(* Logix 5000 project; controller _GigaDiscovery vendor 1 type 14 code 244 rev 35.11; software revision 35.03; part 12 of 23 *)
(* tags used below, declared in another part *)
   LapBars_Alarms_Time : DINT;
   Timer : TIMER[60];
   Timer_Restraints_Open : TIMER[41];
   DC_Field_Motor_7 : UDT_CROUT;   // DC Field Motor 7 Gondola Contactor -Q16101E -Q16103E
   DC_Field_Pylon_Motors : UDT_CROUT;   // DC Field Pylon Motors Contactor -Q10101E -Q10103E
   Emergencies_CL1 : DINT[14];
   Gondola_Drive_Enable : UDT_CROUT;   // Gondola Drive Ch1-Ch2 Start Enable Contactors -Q16105E -Q16107E
   I_EStop_Pb_OCC1 : UDT_DCI_STOP_TEST;   // +OCC E-stop -S30301F
   I_EStop_Pb_OCC2 : UDT_DCI_STOP_TEST;   // +OCC2 E-Stop -S28502F
   I_OCC2_ACONFIRM : BOOL;   // OCC2 Allow Main CONFIRM -S28602F
   I_OCC2_Disable : UDT_DCM;   // OCC 2 CONTROL DISABLE Page 310
   I_OCC2_RESTRAINTS_RELEASE : Sel_3_Pos_2_Input;   // -S28507F RESTRAINTS RELEASE UNLOCK -RUN- LOCK
   I_OCC_Aut_Man_Selector_Motion : UDT_DCM;   // S30801F
   I_OCC_LockOut_Motion : UDT_DCM;   // OCC -Lockout Motion -Q31203E
   I_OCC_Memory_Footpedal : BOOL;
   I_OCC_Temperature_OK : BOOL;   // OCC temperature OK -S31003E
   I_RESTRAINTS_Selector : Sel_3_Pos_2_Input;   // RESTRAINTS Selctor -S30505F Left = Open Right = Close Center = Nothing
   I_Start_PB : Start_AOI;   // Primary console Strat Push botton Right and Left -S30401F -S30403F
   No_Sfty : Std_to_Sfty;
   O_RESTRAINTS_MainValve : UDT_CROUT;   // Main Valve -B40501I
   Power_On_Delay : BOOL;
   Pylon_Start_Drive_1_2 : UDT_CROUT;   // Pylon Start Drive 1 - 2 Contactors -Q9002H -Q9004H -Q10202G
   Pylon_Start_Drive_3_4 : UDT_CROUT;   // Pylon Start Drive 3 - 4 Contactors -Q9005H -Q9007H -Q12202G
   Pylon_Start_Drive_5_6 : UDT_CROUT;   // Pylon Start Drive 5 - 6 Contactors -Q9009E -Q9011E4 -Q14202G -Q14202G
   RESTRAINTS_MainValve_PressTest : Valve_2_pos_monostable;
   RESTRAINTS_Sector : LapBars_Sector[9];
   Start_Stop_Cycle : Sequencer;
(* S_Alarms, continued *)

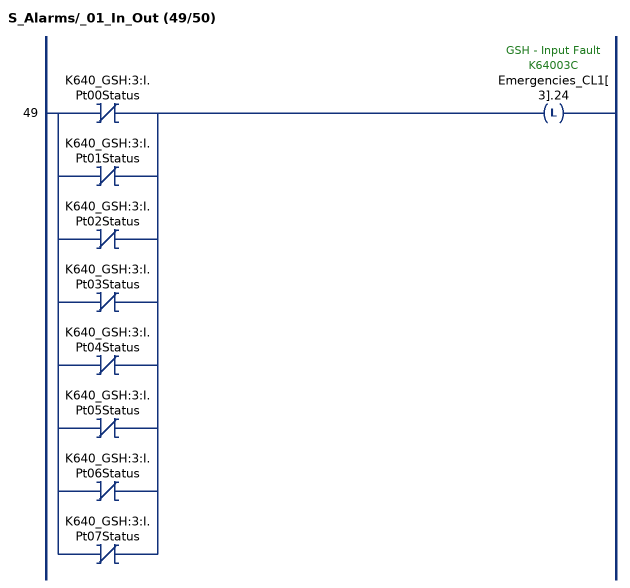
   [picture p209: S_Alarms/_01_In_Out rungs 49-49]
   49: [XIO(K640_GSH:3:I.Pt00Status) ,XIO(K640_GSH:3:I.Pt01Status) ,XIO(K640_GSH:3:I.Pt02Status) ,XIO(K640_GSH:3:I.Pt03Status) ,XIO(K640_GSH:3:I.Pt04Status) ,XIO(K640_GSH:3:I.Pt05Status) ,XIO(K640_GSH:3:I.Pt06Status) ,XIO(K640_GSH:3:I.Pt07Status) ]OTL(Emergencies_CL1[3].24);
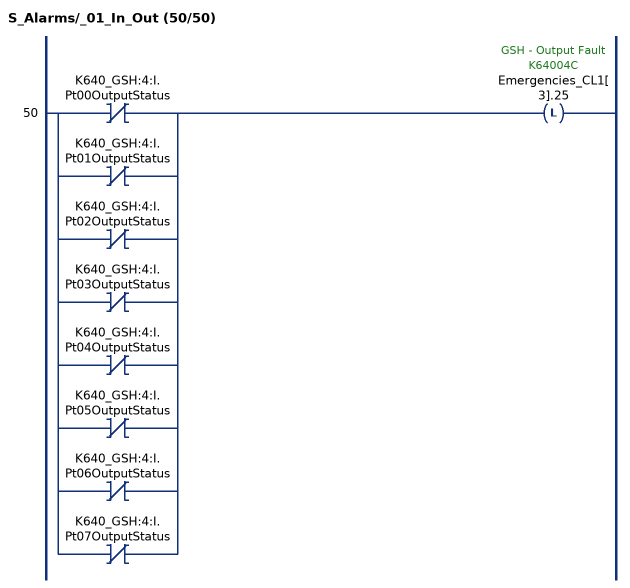
   50: [XIO(K640_GSH:4:I.Pt00OutputStatus) ,XIO(K640_GSH:4:I.Pt01OutputStatus) ,XIO(K640_GSH:4:I.Pt02OutputStatus) ,XIO(K640_GSH:4:I.Pt03OutputStatus) ,XIO(K640_GSH:4:I.Pt04OutputStatus) ,XIO(K640_GSH:4:I.Pt05OutputStatus) ,XIO(K640_GSH:4:I.Pt06OutputStatus) ,XIO(K640_GSH:4:I.Pt07OutputStatus) ]OTL(Emergencies_CL1[3].25);
END_ROUTINE

ROUTINE _02_OCCs   (* ladder *)
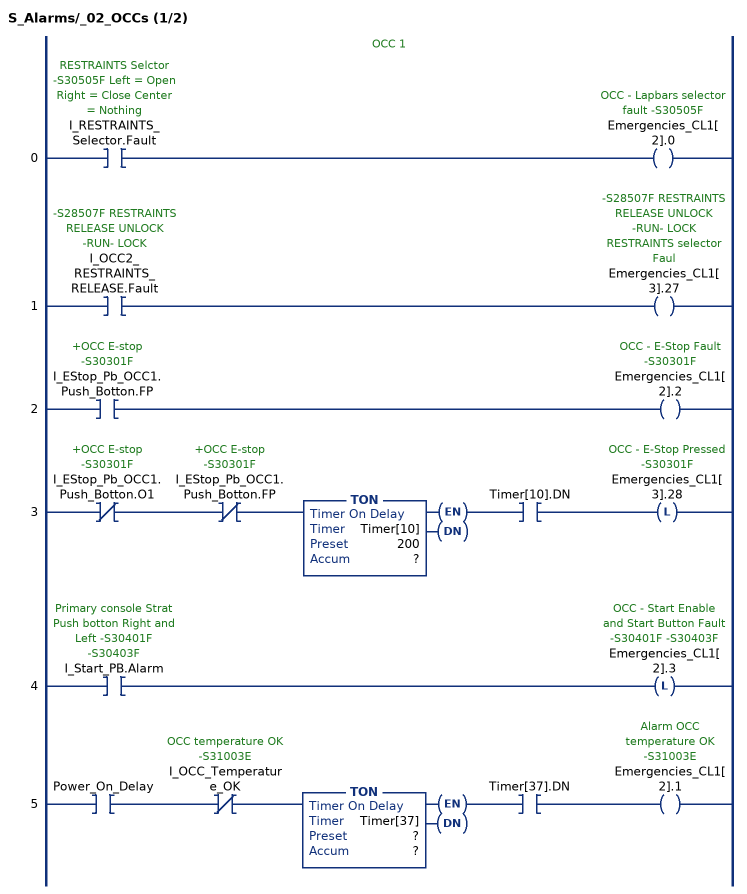
   // OCC 1
   0: XIC(I_RESTRAINTS_Selector.Fault)OTE(Emergencies_CL1[2].0);
   1: XIC(I_OCC2_RESTRAINTS_RELEASE.Fault)OTE(Emergencies_CL1[3].27);
   2: XIC(I_EStop_Pb_OCC1.Push_Botton.FP)OTE(Emergencies_CL1[2].2);
   3: XIO(I_EStop_Pb_OCC1.Push_Botton.O1)XIO(I_EStop_Pb_OCC1.Push_Botton.FP)TON(Timer[10],?,?)XIC(Timer[10].DN)OTL(Emergencies_CL1[3].28);
   4: XIC(I_Start_PB.Alarm)OTL(Emergencies_CL1[2].3);
   5: XIC(Power_On_Delay)XIO(I_OCC_Temperature_OK)TON(Timer[37],?,?)XIC(Timer[37].DN)OTE(Emergencies_CL1[2].1);
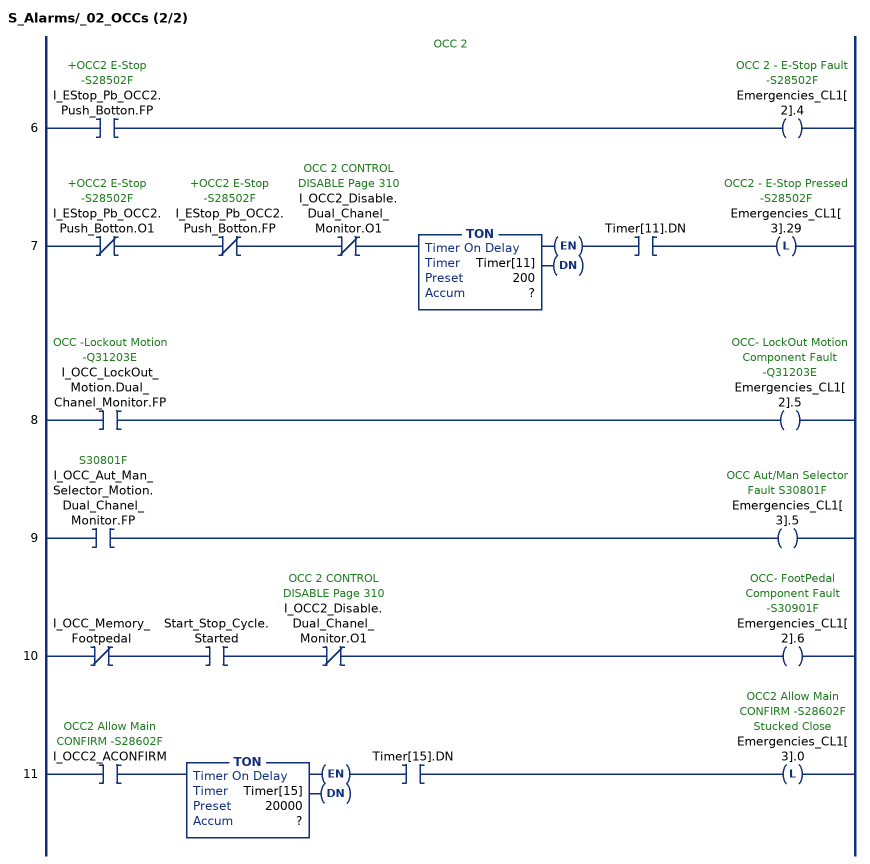
   // OCC 2
   6: XIC(I_EStop_Pb_OCC2.Push_Botton.FP)OTE(Emergencies_CL1[2].4);
   7: XIO(I_EStop_Pb_OCC2.Push_Botton.O1)XIO(I_EStop_Pb_OCC2.Push_Botton.FP)XIO(I_OCC2_Disable.Dual_Chanel_Monitor.O1)TON(Timer[11],?,?)XIC(Timer[11].DN)OTL(Emergencies_CL1[3].29);
   8: XIC(I_OCC_LockOut_Motion.Dual_Chanel_Monitor.FP)OTE(Emergencies_CL1[2].5);
   9: XIC(I_OCC_Aut_Man_Selector_Motion.Dual_Chanel_Monitor.FP)OTE(Emergencies_CL1[3].5);
   10: XIO(I_OCC_Memory_Footpedal)XIC(Start_Stop_Cycle.Started)XIO(I_OCC2_Disable.Dual_Chanel_Monitor.O1)OTE(Emergencies_CL1[2].6);
   11: XIC(I_OCC2_ACONFIRM)TON(Timer[15],?,?)XIC(Timer[15].DN)OTL(Emergencies_CL1[3].0);
END_ROUTINE

ROUTINE _03_MCC   (* ladder *)
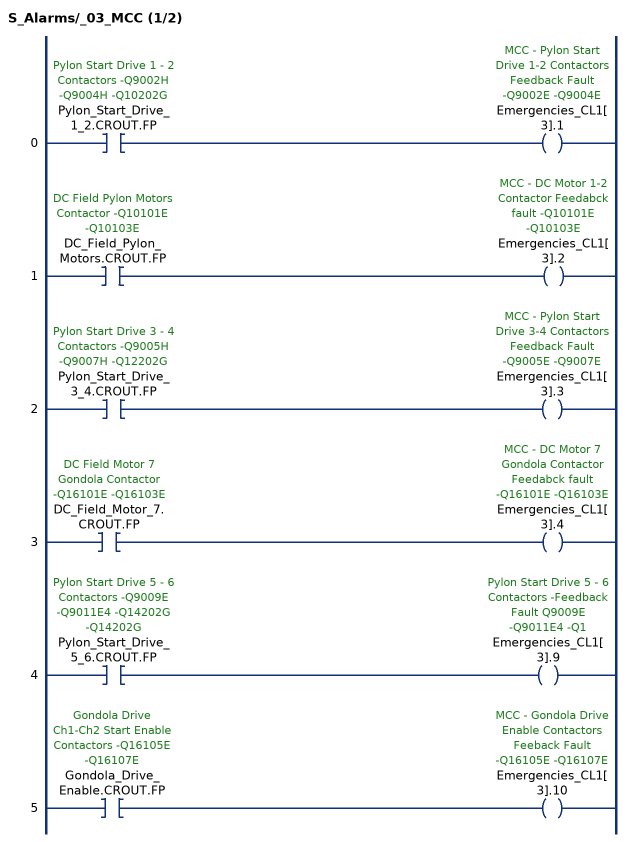
   0: XIC(Pylon_Start_Drive_1_2.CROUT.FP)OTE(Emergencies_CL1[3].1);
   1: XIC(DC_Field_Pylon_Motors.CROUT.FP)OTE(Emergencies_CL1[3].2);
   2: XIC(Pylon_Start_Drive_3_4.CROUT.FP)OTE(Emergencies_CL1[3].3);
   3: XIC(DC_Field_Motor_7.CROUT.FP)OTE(Emergencies_CL1[3].4);
   4: XIC(Pylon_Start_Drive_5_6.CROUT.FP)OTE(Emergencies_CL1[3].9);
   5: XIC(Gondola_Drive_Enable.CROUT.FP)OTE(Emergencies_CL1[3].10);
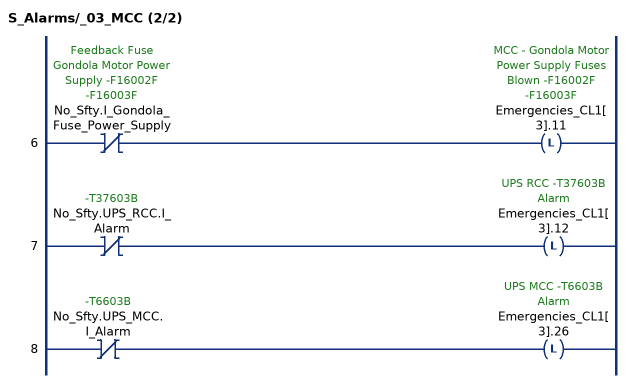
   6: XIO(No_Sfty.I_Gondola_Fuse_Power_Supply)OTL(Emergencies_CL1[3].11);
   7: XIO(No_Sfty.UPS_RCC.I_Alarm)OTL(Emergencies_CL1[3].12);
   8: XIO(No_Sfty.UPS_MCC.I_Alarm)OTL(Emergencies_CL1[3].26);
END_ROUTINE

ROUTINE _04_RESTRAINT_RELEASE   (* ladder *)
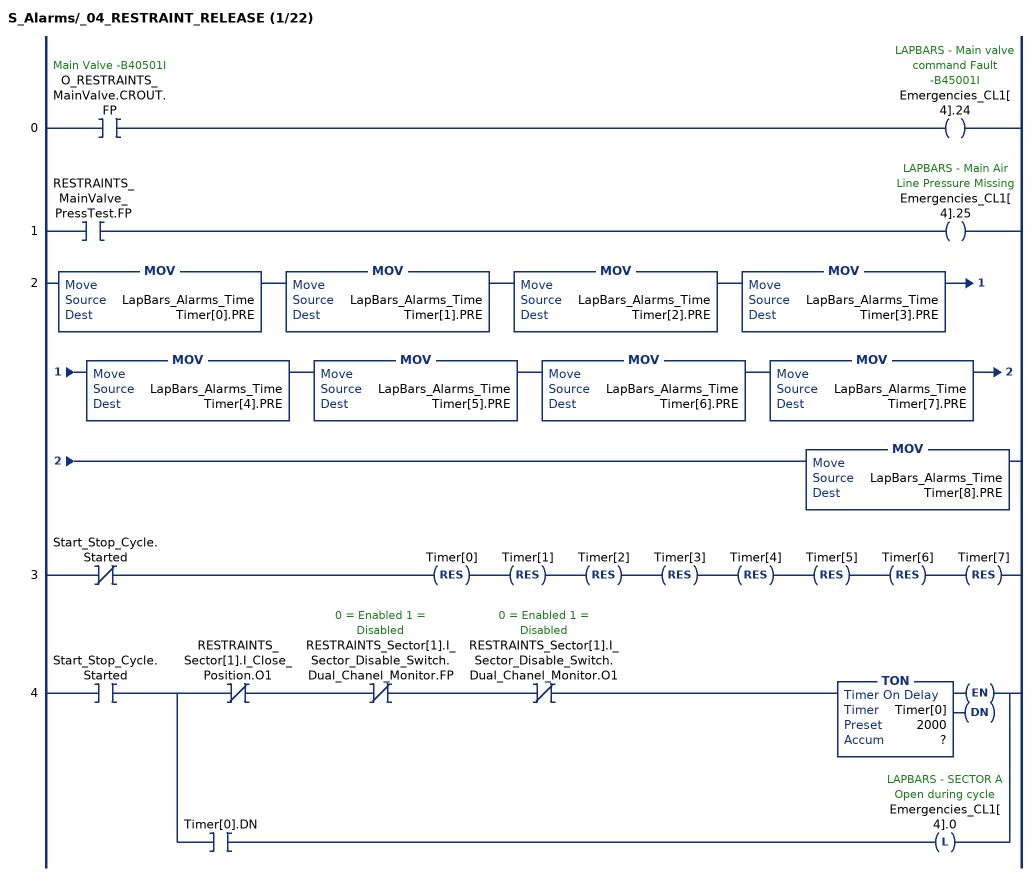
   0: XIC(O_RESTRAINTS_MainValve.CROUT.FP)OTE(Emergencies_CL1[4].24);
   1: XIC(RESTRAINTS_MainValve_PressTest.FP)OTE(Emergencies_CL1[4].25);
   2: MOV(LapBars_Alarms_Time,Timer[0].PRE)MOV(LapBars_Alarms_Time,Timer[1].PRE)MOV(LapBars_Alarms_Time,Timer[2].PRE)MOV(LapBars_Alarms_Time,Timer[3].PRE)MOV(LapBars_Alarms_Time,Timer[4].PRE)MOV(LapBars_Alarms_Time,Timer[5].PRE)MOV(LapBars_Alarms_Time,Timer[6].PRE)MOV(LapBars_Alarms_Time,Timer[7].PRE)MOV(LapBars_Alarms_Time,Timer[8].PRE);
   3: XIO(Start_Stop_Cycle.Started)RES(Timer[0])RES(Timer[1])RES(Timer[2])RES(Timer[3])RES(Timer[4])RES(Timer[5])RES(Timer[6])RES(Timer[7]);
   4: XIC(Start_Stop_Cycle.Started)[XIO(RESTRAINTS_Sector[1].I_Close_Position.O1) XIO(RESTRAINTS_Sector[1].I_Sector_Disable_Switch.Dual_Chanel_Monitor.FP) XIO(RESTRAINTS_Sector[1].I_Sector_Disable_Switch.Dual_Chanel_Monitor.O1) TON(Timer[0],?,?) ,XIC(Timer[0].DN) OTL(Emergencies_CL1[4].0) ];
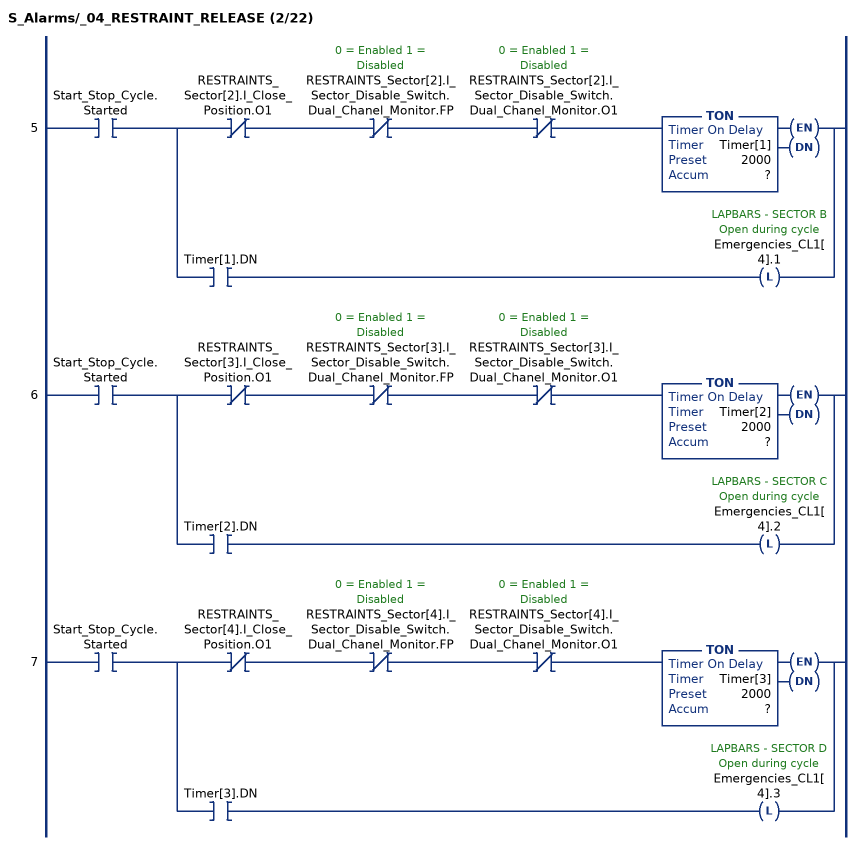
   5: XIC(Start_Stop_Cycle.Started)[XIO(RESTRAINTS_Sector[2].I_Close_Position.O1) XIO(RESTRAINTS_Sector[2].I_Sector_Disable_Switch.Dual_Chanel_Monitor.FP) XIO(RESTRAINTS_Sector[2].I_Sector_Disable_Switch.Dual_Chanel_Monitor.O1) TON(Timer[1],?,?) ,XIC(Timer[1].DN) OTL(Emergencies_CL1[4].1) ];
   6: XIC(Start_Stop_Cycle.Started)[XIO(RESTRAINTS_Sector[3].I_Close_Position.O1) XIO(RESTRAINTS_Sector[3].I_Sector_Disable_Switch.Dual_Chanel_Monitor.FP) XIO(RESTRAINTS_Sector[3].I_Sector_Disable_Switch.Dual_Chanel_Monitor.O1) TON(Timer[2],?,?) ,XIC(Timer[2].DN) OTL(Emergencies_CL1[4].2) ];
   7: XIC(Start_Stop_Cycle.Started)[XIO(RESTRAINTS_Sector[4].I_Close_Position.O1) XIO(RESTRAINTS_Sector[4].I_Sector_Disable_Switch.Dual_Chanel_Monitor.FP) XIO(RESTRAINTS_Sector[4].I_Sector_Disable_Switch.Dual_Chanel_Monitor.O1) TON(Timer[3],?,?) ,XIC(Timer[3].DN) OTL(Emergencies_CL1[4].3) ];
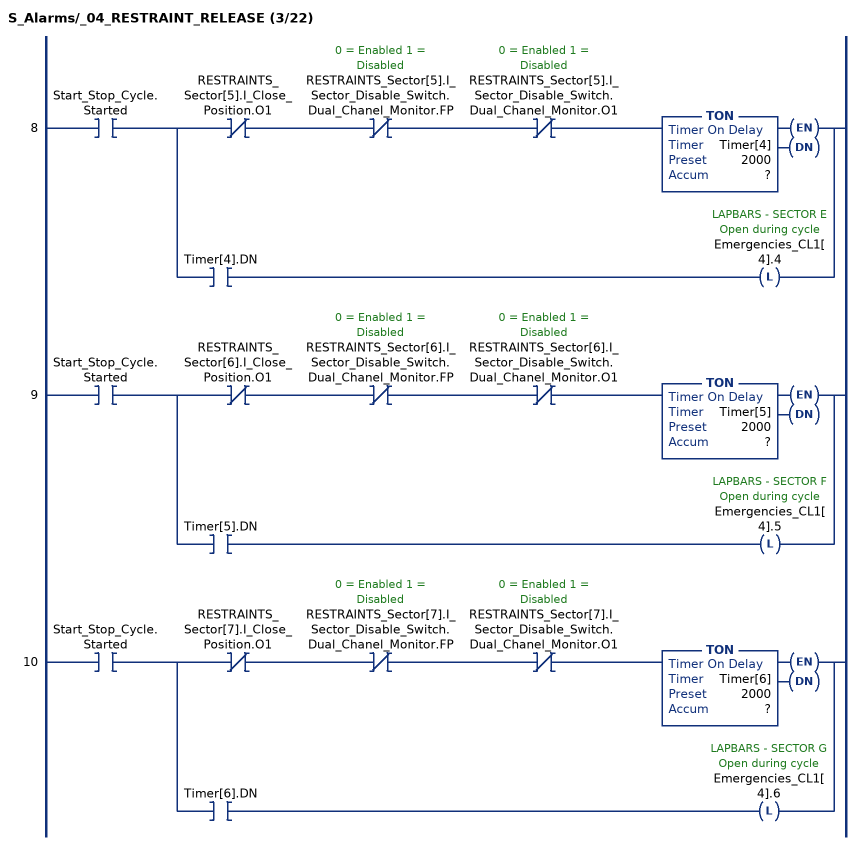
   8: XIC(Start_Stop_Cycle.Started)[XIO(RESTRAINTS_Sector[5].I_Close_Position.O1) XIO(RESTRAINTS_Sector[5].I_Sector_Disable_Switch.Dual_Chanel_Monitor.FP) XIO(RESTRAINTS_Sector[5].I_Sector_Disable_Switch.Dual_Chanel_Monitor.O1) TON(Timer[4],?,?) ,XIC(Timer[4].DN) OTL(Emergencies_CL1[4].4) ];
   9: XIC(Start_Stop_Cycle.Started)[XIO(RESTRAINTS_Sector[6].I_Close_Position.O1) XIO(RESTRAINTS_Sector[6].I_Sector_Disable_Switch.Dual_Chanel_Monitor.FP) XIO(RESTRAINTS_Sector[6].I_Sector_Disable_Switch.Dual_Chanel_Monitor.O1) TON(Timer[5],?,?) ,XIC(Timer[5].DN) OTL(Emergencies_CL1[4].5) ];
   10: XIC(Start_Stop_Cycle.Started)[XIO(RESTRAINTS_Sector[7].I_Close_Position.O1) XIO(RESTRAINTS_Sector[7].I_Sector_Disable_Switch.Dual_Chanel_Monitor.FP) XIO(RESTRAINTS_Sector[7].I_Sector_Disable_Switch.Dual_Chanel_Monitor.O1) TON(Timer[6],?,?) ,XIC(Timer[6].DN) OTL(Emergencies_CL1[4].6) ];
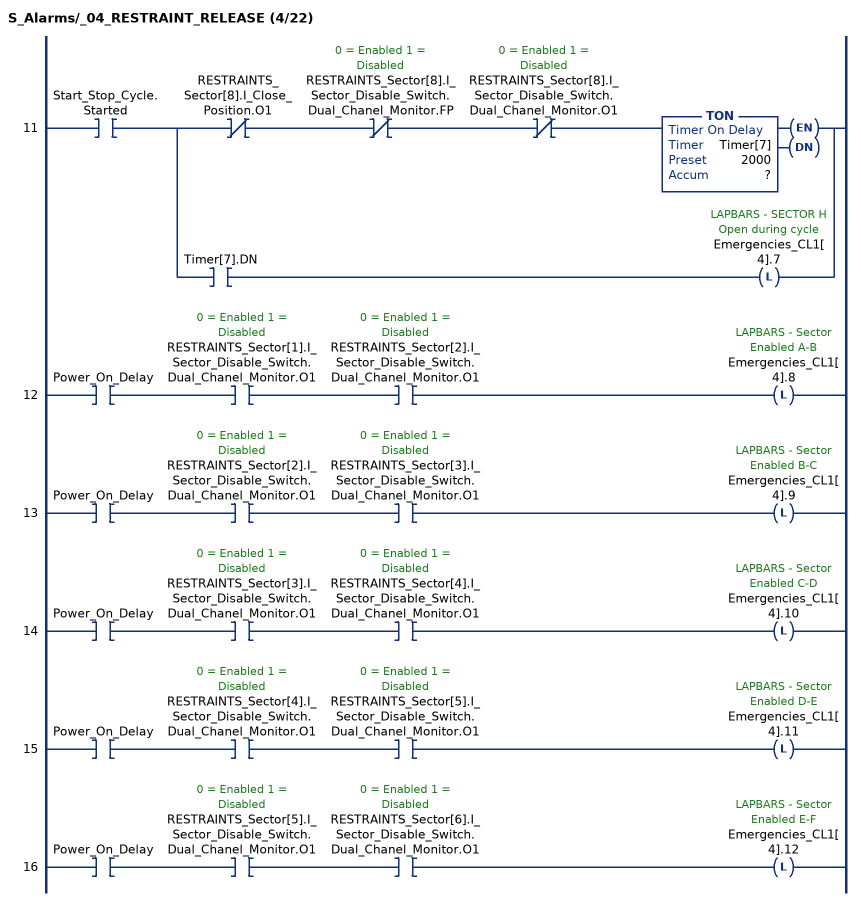
   11: XIC(Start_Stop_Cycle.Started)[XIO(RESTRAINTS_Sector[8].I_Close_Position.O1) XIO(RESTRAINTS_Sector[8].I_Sector_Disable_Switch.Dual_Chanel_Monitor.FP) XIO(RESTRAINTS_Sector[8].I_Sector_Disable_Switch.Dual_Chanel_Monitor.O1) TON(Timer[7],?,?) ,XIC(Timer[7].DN) OTL(Emergencies_CL1[4].7) ];
   12: XIC(Power_On_Delay)XIC(RESTRAINTS_Sector[1].I_Sector_Disable_Switch.Dual_Chanel_Monitor.O1)XIC(RESTRAINTS_Sector[2].I_Sector_Disable_Switch.Dual_Chanel_Monitor.O1)OTL(Emergencies_CL1[4].8);
   13: XIC(Power_On_Delay)XIC(RESTRAINTS_Sector[2].I_Sector_Disable_Switch.Dual_Chanel_Monitor.O1)XIC(RESTRAINTS_Sector[3].I_Sector_Disable_Switch.Dual_Chanel_Monitor.O1)OTL(Emergencies_CL1[4].9);
   14: XIC(Power_On_Delay)XIC(RESTRAINTS_Sector[3].I_Sector_Disable_Switch.Dual_Chanel_Monitor.O1)XIC(RESTRAINTS_Sector[4].I_Sector_Disable_Switch.Dual_Chanel_Monitor.O1)OTL(Emergencies_CL1[4].10);
   15: XIC(Power_On_Delay)XIC(RESTRAINTS_Sector[4].I_Sector_Disable_Switch.Dual_Chanel_Monitor.O1)XIC(RESTRAINTS_Sector[5].I_Sector_Disable_Switch.Dual_Chanel_Monitor.O1)OTL(Emergencies_CL1[4].11);
   16: XIC(Power_On_Delay)XIC(RESTRAINTS_Sector[5].I_Sector_Disable_Switch.Dual_Chanel_Monitor.O1)XIC(RESTRAINTS_Sector[6].I_Sector_Disable_Switch.Dual_Chanel_Monitor.O1)OTL(Emergencies_CL1[4].12);
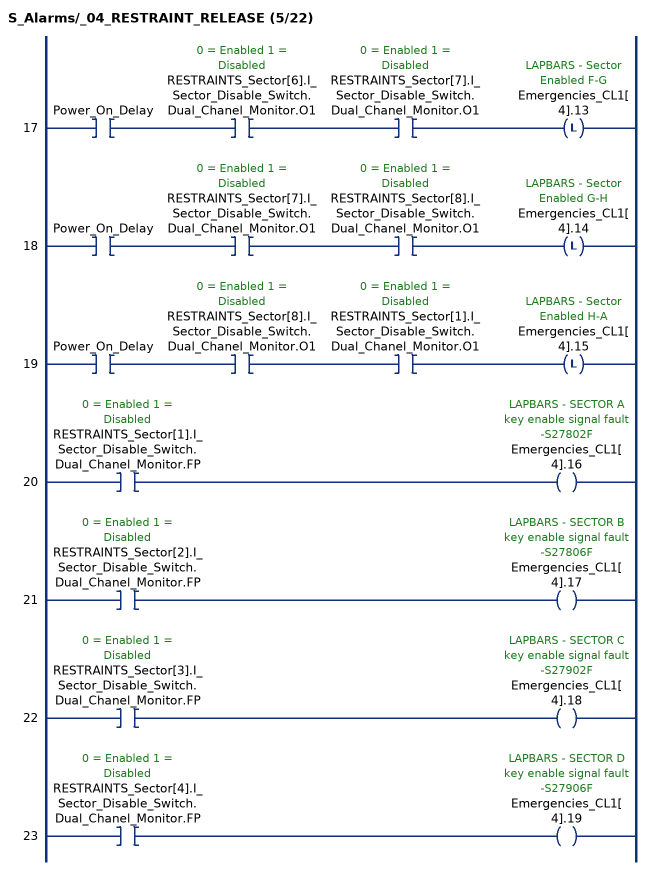
   17: XIC(Power_On_Delay)XIC(RESTRAINTS_Sector[6].I_Sector_Disable_Switch.Dual_Chanel_Monitor.O1)XIC(RESTRAINTS_Sector[7].I_Sector_Disable_Switch.Dual_Chanel_Monitor.O1)OTL(Emergencies_CL1[4].13);
   18: XIC(Power_On_Delay)XIC(RESTRAINTS_Sector[7].I_Sector_Disable_Switch.Dual_Chanel_Monitor.O1)XIC(RESTRAINTS_Sector[8].I_Sector_Disable_Switch.Dual_Chanel_Monitor.O1)OTL(Emergencies_CL1[4].14);
   19: XIC(Power_On_Delay)XIC(RESTRAINTS_Sector[8].I_Sector_Disable_Switch.Dual_Chanel_Monitor.O1)XIC(RESTRAINTS_Sector[1].I_Sector_Disable_Switch.Dual_Chanel_Monitor.O1)OTL(Emergencies_CL1[4].15);
   20: XIC(RESTRAINTS_Sector[1].I_Sector_Disable_Switch.Dual_Chanel_Monitor.FP)OTE(Emergencies_CL1[4].16);
   21: XIC(RESTRAINTS_Sector[2].I_Sector_Disable_Switch.Dual_Chanel_Monitor.FP)OTE(Emergencies_CL1[4].17);
   22: XIC(RESTRAINTS_Sector[3].I_Sector_Disable_Switch.Dual_Chanel_Monitor.FP)OTE(Emergencies_CL1[4].18);
   23: XIC(RESTRAINTS_Sector[4].I_Sector_Disable_Switch.Dual_Chanel_Monitor.FP)OTE(Emergencies_CL1[4].19);
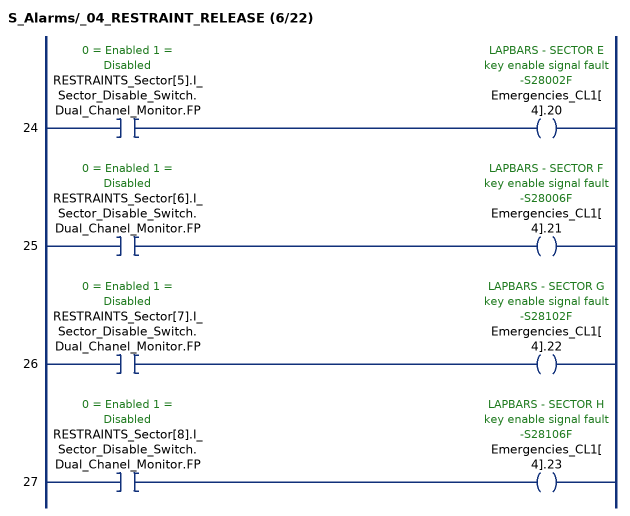
   24: XIC(RESTRAINTS_Sector[5].I_Sector_Disable_Switch.Dual_Chanel_Monitor.FP)OTE(Emergencies_CL1[4].20);
   25: XIC(RESTRAINTS_Sector[6].I_Sector_Disable_Switch.Dual_Chanel_Monitor.FP)OTE(Emergencies_CL1[4].21);
   26: XIC(RESTRAINTS_Sector[7].I_Sector_Disable_Switch.Dual_Chanel_Monitor.FP)OTE(Emergencies_CL1[4].22);
   27: XIC(RESTRAINTS_Sector[8].I_Sector_Disable_Switch.Dual_Chanel_Monitor.FP)OTE(Emergencies_CL1[4].23);
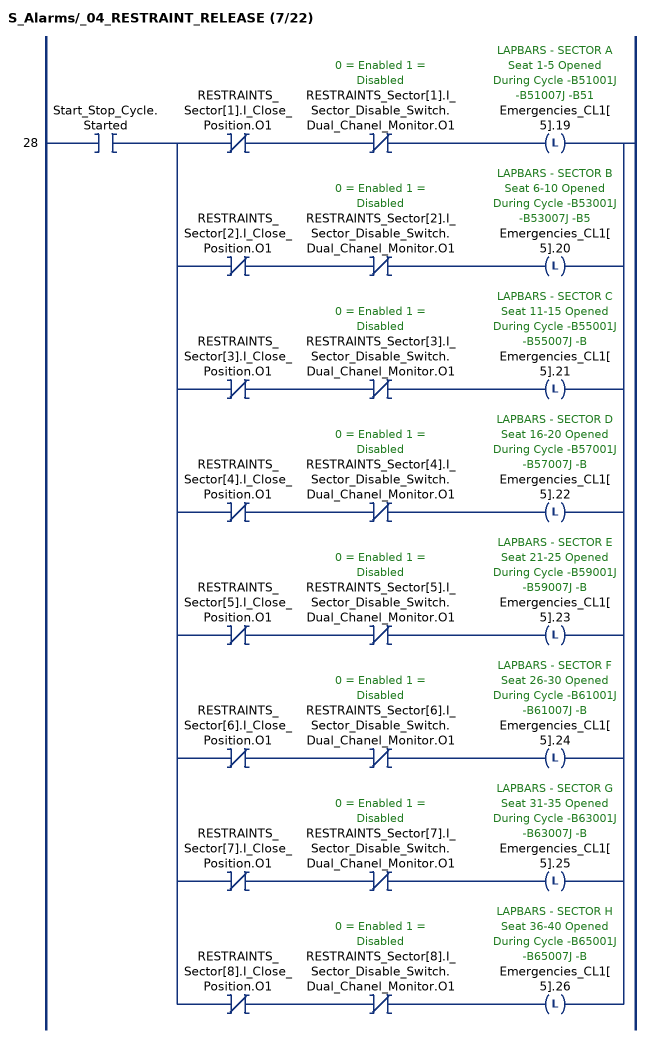
   28: XIC(Start_Stop_Cycle.Started)[XIO(RESTRAINTS_Sector[1].I_Close_Position.O1) XIO(RESTRAINTS_Sector[1].I_Sector_Disable_Switch.Dual_Chanel_Monitor.O1) OTL(Emergencies_CL1[5].19) ,XIO(RESTRAINTS_Sector[2].I_Close_Position.O1) XIO(RESTRAINTS_Sector[2].I_Sector_Disable_Switch.Dual_Chanel_Monitor.O1) OTL(Emergencies_CL1[5].20) ,XIO(RESTRAINTS_Sector[3].I_Close_Position.O1) XIO(RESTRAINTS_Sector[3].I_Sector_Disable_Switch.Dual_Chanel_Monitor.O1) OTL(Emergencies_CL1[5].21) ,XIO(RESTRAINTS_Sector[4].I_Close_Position.O1) XIO(RESTRAINTS_Sector[4].I_Sector_Disable_Switch.Dual_Chanel_Monitor.O1) OTL(Emergencies_CL1[5].22) ,XIO(RESTRAINTS_Sector[5].I_Close_Position.O1) XIO(RESTRAINTS_Sector[5].I_Sector_Disable_Switch.Dual_Chanel_Monitor.O1) OTL(Emergencies_CL1[5].23) ,XIO(RESTRAINTS_Sector[6].I_Close_Position.O1) XIO(RESTRAINTS_Sector[6].I_Sector_Disable_Switch.Dual_Chanel_Monitor.O1) OTL(Emergencies_CL1[5].24) ,XIO(RESTRAINTS_Sector[7].I_Close_Position.O1) XIO(RESTRAINTS_Sector[7].I_Sector_Disable_Switch.Dual_Chanel_Monitor.O1) OTL(Emergencies_CL1[5].25) ,XIO(RESTRAINTS_Sector[8].I_Close_Position.O1) XIO(RESTRAINTS_Sector[8].I_Sector_Disable_Switch.Dual_Chanel_Monitor.O1) OTL(Emergencies_CL1[5].26) ];